screen "0887_Create Part Counter" 1280x800, template "Navigation"
   on GenerateScreen: SetTag("Create Part Counter Control", 1); SetTag("Create Part Counter Multiplexing Control", 0); function_b431313b("Part Counter Name", U 1, N)
   TextField "Text field_1" at 137,226 size 48x32; Text '1.'
      Visibility <- "Create Part Counter Control"
   TextField "Text field_2" at 137,266 size 48x32; Text '2.'
      Visibility <- "Create Part Counter Control"
   TextField "Text field_3" at 137,306 size 48x32; Text '3.'
      Visibility <- "Create Part Counter Control"
   TextField "Text field_4" at 137,346 size 48x32; Text '4.'
      Visibility <- "Create Part Counter Control"
   TextField "Text field_5" at 137,386 size 48x32; Text '5.'
      Visibility <- "Create Part Counter Control"
   TextField "Text field_6" at 137,426 size 48x32; Text '6.'
      Visibility <- "Create Part Counter Control"
   TextField "Text field_7" at 137,466 size 48x32; Text '7.'
      Visibility <- "Create Part Counter Control"
   TextField "Text field_8" at 137,506 size 48x32; Text '8.'
      Visibility <- "Create Part Counter Control"
   TextField "Text field_9" at 137,546 size 48x32; Text '9.'
      Visibility <- "Create Part Counter Control"
   TextField "Text field_10" at 137,586 size 48x32; Text '10.'
      Visibility <- "Create Part Counter Control"
   TextField "Text field_11" at 489,226 size 48x32; Text '11.'
      Visibility <- "Create Part Counter Control"
   TextField "Text field_12" at 489,266 size 48x32; Text '12.'
      Visibility <- "Create Part Counter Control"
   TextField "Text field_13" at 489,306 size 48x32; Text '13.'
      Visibility <- "Create Part Counter Control"
   TextField "Text field_14" at 489,346 size 48x32; Text '14.'
      Visibility <- "Create Part Counter Control"
   TextField "Text field_15" at 489,386 size 48x32; Text '15.'
      Visibility <- "Create Part Counter Control"
   TextField "Text field_16" at 489,426 size 48x32; Text '16.'
      Visibility <- "Create Part Counter Control"
   TextField "Text field_17" at 489,466 size 48x32; Text '17.'
      Visibility <- "Create Part Counter Control"
   TextField "Text field_18" at 489,506 size 48x32; Text '18.'
      Visibility <- "Create Part Counter Control"
   TextField "Text field_19" at 489,546 size 48x32; Text '19.'
      Visibility <- "Create Part Counter Control"
   TextField "Text field_20" at 489,586 size 48x32; Text '20.'
      Visibility <- "Create Part Counter Control"
   TextField "Text field_21" at 832,226 size 48x32; Text '21.'
      Visibility <- "Create Part Counter Control"
   TextField "Text field_22" at 832,266 size 48x32; Text '22.'
      Visibility <- "Create Part Counter Control"
   TextField "Text field_23" at 832,306 size 48x32; Text '23.'
      Visibility <- "Create Part Counter Control"
   TextField "Text field_24" at 832,346 size 48x32; Text '24.'
      Visibility <- "Create Part Counter Control"
   TextField "Text field_25" at 832,386 size 48x32; Text '25.'
      Visibility <- "Create Part Counter Control"
   TextField "Text field_26" at 832,426 size 48x32; Text '26.'
      Visibility <- "Create Part Counter Control"
   TextField "Text field_27" at 832,466 size 48x32; Text '27.'
      Visibility <- "Create Part Counter Control"
   TextField "Text field_28" at 832,506 size 48x32; Text '28.'
      Visibility <- "Create Part Counter Control"
   TextField "Text field_29" at 832,546 size 48x32; Text '29.'
      Visibility <- "Create Part Counter Control"
   TextField "Text field_30" at 832,586 size 48x32; Text '30.'
      Visibility <- "Create Part Counter Control"
   TextField "Text field_31" at 137,226 size 48x32; Text '31.'
      Visibility <- "Create Part Counter Control"
   TextField "Text field_32" at 137,266 size 48x32; Text '32.'
      Visibility <- "Create Part Counter Control"
   TextField "Text field_33" at 137,306 size 48x32; Text '33.'
      Visibility <- "Create Part Counter Control"
   TextField "Text field_34" at 137,346 size 48x32; Text '34.'
      Visibility <- "Create Part Counter Control"
   TextField "Text field_35" at 137,386 size 48x32; Text '35.'
      Visibility <- "Create Part Counter Control"
   TextField "Text field_36" at 137,426 size 48x32; Text '36.'
      Visibility <- "Create Part Counter Control"
   TextField "Text field_37" at 137,466 size 48x32; Text '37.'
      Visibility <- "Create Part Counter Control"
   TextField "Text field_38" at 137,506 size 48x32; Text '38.'
      Visibility <- "Create Part Counter Control"
   TextField "Text field_39" at 137,546 size 48x32; Text '39.'
      Visibility <- "Create Part Counter Control"
   TextField "Text field_40" at 137,586 size 48x32; Text '40.'
      Visibility <- "Create Part Counter Control"
   TextField "Text field_41" at 489,226 size 48x32; Text '41.'
      Visibility <- "Create Part Counter Control"
   TextField "Text field_42" at 489,266 size 48x32; Text '42.'
      Visibility <- "Create Part Counter Control"
   TextField "Text field_43" at 489,306 size 48x32; Text '43.'
      Visibility <- "Create Part Counter Control"
   TextField "Text field_44" at 489,346 size 48x32; Text '44.'
      Visibility <- "Create Part Counter Control"
   TextField "Text field_45" at 489,386 size 48x32; Text '45.'
      Visibility <- "Create Part Counter Control"
   TextField "Text field_46" at 489,426 size 48x32; Text '46.'
      Visibility <- "Create Part Counter Control"
   TextField "Text field_47" at 489,466 size 48x32; Text '47.'
      Visibility <- "Create Part Counter Control"
   TextField "Text field_48" at 489,506 size 48x32; Text '48.'
      Visibility <- "Create Part Counter Control"
   TextField "Text field_49" at 489,546 size 48x32; Text '49.'
      Visibility <- "Create Part Counter Control"
   TextField "Text field_50" at 489,586 size 48x32; Text '50.'
      Visibility <- "Create Part Counter Control"
   TextField "Text field_51" at 832,226 size 48x32; Text '51.'
      Visibility <- "Create Part Counter Control"
   TextField "Text field_52" at 832,266 size 48x32; Text '52.'
      Visibility <- "Create Part Counter Control"
   TextField "Text field_53" at 832,306 size 48x32; Text '53.'
      Visibility <- "Create Part Counter Control"
   TextField "Text field_54" at 832,346 size 48x32; Text '54.'
      Visibility <- "Create Part Counter Control"
   TextField "Text field_55" at 832,386 size 48x32; Text '55.'
      Visibility <- "Create Part Counter Control"
   TextField "Text field_56" at 832,426 size 48x32; Text '56.'
      Visibility <- "Create Part Counter Control"
   TextField "Text field_57" at 832,466 size 48x32; Text '57.'
      Visibility <- "Create Part Counter Control"
   TextField "Text field_58" at 832,506 size 48x32; Text '58.'
      Visibility <- "Create Part Counter Control"
   TextField "Text field_59" at 832,546 size 48x32; Text '59.'
      Visibility <- "Create Part Counter Control"
   TextField "Text field_60" at 832,586 size 48x32; Text '60.'
      Visibility <- "Create Part Counter Control"
   TextField "Text field_61" at 137,226 size 48x32; Text '61.'
      Visibility <- "Create Part Counter Control"
   TextField "Text field_62" at 137,266 size 48x32; Text '62.'
      Visibility <- "Create Part Counter Control"
   TextField "Text field_63" at 137,306 size 48x32; Text '63.'
      Visibility <- "Create Part Counter Control"
   TextField "Text field_64" at 137,346 size 48x32; Text '64.'
      Visibility <- "Create Part Counter Control"
   TextField "Text field_65" at 137,386 size 48x32; Text '65.'
      Visibility <- "Create Part Counter Control"
   TextField "Text field_66" at 137,426 size 48x32; Text '66.'
      Visibility <- "Create Part Counter Control"
   TextField "Text field_67" at 137,466 size 48x32; Text '67.'
      Visibility <- "Create Part Counter Control"
   TextField "Text field_68" at 137,506 size 48x32; Text '68.'
      Visibility <- "Create Part Counter Control"
   TextField "Text field_69" at 137,546 size 48x32; Text '69.'
      Visibility <- "Create Part Counter Control"
   TextField "Text field_70" at 137,586 size 48x32; Text '70.'
      Visibility <- "Create Part Counter Control"
   TextField "Text field_71" at 489,226 size 48x32; Text '71.'
      Visibility <- "Create Part Counter Control"
   TextField "Text field_72" at 489,266 size 48x32; Text '72.'
      Visibility <- "Create Part Counter Control"
   TextField "Text field_73" at 489,306 size 48x32; Text '73.'
      Visibility <- "Create Part Counter Control"
   TextField "Text field_74" at 489,346 size 48x32; Text '74.'
      Visibility <- "Create Part Counter Control"
   TextField "Text field_75" at 489,386 size 48x32; Text '75.'
      Visibility <- "Create Part Counter Control"
   TextField "Text field_76" at 489,426 size 48x32; Text '76.'
      Visibility <- "Create Part Counter Control"
   TextField "Text field_77" at 489,466 size 48x32; Text '77.'
      Visibility <- "Create Part Counter Control"
   TextField "Text field_78" at 489,506 size 48x32; Text '78.'
      Visibility <- "Create Part Counter Control"
   TextField "Text field_79" at 489,546 size 48x32; Text '79.'
      Visibility <- "Create Part Counter Control"
   TextField "Text field_80" at 489,586 size 48x32; Text '80.'
      Visibility <- "Create Part Counter Control"
   TextField "Text field_81" at 832,226 size 48x32; Text '81.'
      Visibility <- "Create Part Counter Control"
   TextField "Text field_82" at 832,266 size 48x32; Text '82.'
      Visibility <- "Create Part Counter Control"
   TextField "Text field_83" at 832,306 size 48x32; Text '83.'
      Visibility <- "Create Part Counter Control"
   TextField "Text field_84" at 832,346 size 48x32; Text '84.'
      Visibility <- "Create Part Counter Control"
   TextField "Text field_85" at 832,386 size 48x32; Text '85.'
      Visibility <- "Create Part Counter Control"
   TextField "Text field_86" at 832,426 size 48x32; Text '86.'
      Visibility <- "Create Part Counter Control"
   TextField "Text field_87" at 832,466 size 48x32; Text '87.'
      Visibility <- "Create Part Counter Control"
   TextField "Text field_88" at 832,506 size 48x32; Text '88.'
      Visibility <- "Create Part Counter Control"
   TextField "Text field_89" at 832,546 size 48x32; Text '89.'
      Visibility <- "Create Part Counter Control"
   TextField "Text field_90" at 832,586 size 48x32; Text '90.'
      Visibility <- "Create Part Counter Control"
   TextField "Text field_151" at 489,226 size 48x32; Text '101.'
      Visibility <- "Create Part Counter Control"
   TextField "Text field_152" at 489,266 size 48x32; Text '102.'
      Visibility <- "Create Part Counter Control"
   TextField "Text field_153" at 489,306 size 48x32; Text '103.'
      Visibility <- "Create Part Counter Control"
   TextField "Text field_154" at 489,346 size 48x32; Text '104.'
      Visibility <- "Create Part Counter Control"
   TextField "Text field_155" at 489,386 size 48x32; Text '105.'
      Visibility <- "Create Part Counter Control"
   TextField "Text field_156" at 489,426 size 48x32; Text '106.'
      Visibility <- "Create Part Counter Control"
   TextField "Text field_157" at 489,466 size 48x32; Text '107.'
      Visibility <- "Create Part Counter Control"
   TextField "Text field_158" at 489,506 size 48x32; Text '108.'
      Visibility <- "Create Part Counter Control"
   TextField "Text field_159" at 489,546 size 48x32; Text '109.'
      Visibility <- "Create Part Counter Control"
   TextField "Text field_160" at 489,586 size 48x32; Text '110.'
      Visibility <- "Create Part Counter Control"
   TextField "Text field_161" at 832,226 size 48x32; Text '111.'
      Visibility <- "Create Part Counter Control"
   TextField "Text field_162" at 832,266 size 48x32; Text '112.'
      Visibility <- "Create Part Counter Control"
   TextField "Text field_163" at 832,306 size 48x32; Text '113.'
      Visibility <- "Create Part Counter Control"
   TextField "Text field_164" at 832,346 size 48x32; Text '114.'
      Visibility <- "Create Part Counter Control"
   TextField "Text field_165" at 832,386 size 48x32; Text '115.'
      Visibility <- "Create Part Counter Control"
   TextField "Text field_166" at 832,426 size 48x32; Text '116.'
      Visibility <- "Create Part Counter Control"
   TextField "Text field_167" at 832,466 size 48x32; Text '117.'
      Visibility <- "Create Part Counter Control"
   TextField "Text field_168" at 832,506 size 48x32; Text '118.'
      Visibility <- "Create Part Counter Control"
   TextField "Text field_169" at 832,546 size 48x32; Text '119.'
      Visibility <- "Create Part Counter Control"
   TextField "Text field_170" at 832,586 size 48x32; Text '120.'
      Visibility <- "Create Part Counter Control"
   TextField "Text field_171" at 137,226 size 48x32; Text '91.'
      Visibility <- "Create Part Counter Control"
   TextField "Text field_172" at 137,266 size 48x32; Text '92.'
      Visibility <- "Create Part Counter Control"
   TextField "Text field_173" at 137,306 size 48x32; Text '93.'
      Visibility <- "Create Part Counter Control"
   TextField "Text field_174" at 137,346 size 48x32; Text '94.'
      Visibility <- "Create Part Counter Control"
   TextField "Text field_175" at 137,386 size 48x32; Text '95.'
      Visibility <- "Create Part Counter Control"
   TextField "Text field_176" at 137,426 size 48x32; Text '96.'
      Visibility <- "Create Part Counter Control"
   TextField "Text field_177" at 137,466 size 48x32; Text '97.'
      Visibility <- "Create Part Counter Control"
   TextField "Text field_178" at 137,506 size 48x32; Text '98.'
      Visibility <- "Create Part Counter Control"
   TextField "Text field_179" at 137,546 size 48x32; Text '99.'
      Visibility <- "Create Part Counter Control"
   TextField "Text field_180" at 137,586 size 48x32; Text '100.'
      Visibility <- "Create Part Counter Control"
   IOField "NamePart1" at 207,225 size 240x32; FormatPattern ????????????????????
      on OnFinishInput: SetTag("Create Part Counter Button Save", 1)
      ProcessValue <- "Part_Counter_Coloum_1"
   Button "Button_3" at 326,104 size 451x32; TextOff 'Create Part Counter'
   IOField "NamePart2" at 207,265 size 240x32; FormatPattern ????????????????????
      on OnFinishInput: SetTag("Create Part Counter Button Save", 1)
      ProcessValue <- "Part_Counter_Coloum_2"
   IOField "NamePart3" at 207,305 size 240x32; FormatPattern ????????????????????
      on OnFinishInput: SetTag("Create Part Counter Button Save", 1)
      ProcessValue <- "Part_Counter_Coloum_3"
   IOField "NamePart4" at 207,345 size 240x32; FormatPattern ????????????????????
      on OnFinishInput: SetTag("Create Part Counter Button Save", 1)
      ProcessValue <- "Part_Counter_Coloum_4"
   IOField "NamePart5" at 207,385 size 240x32; FormatPattern ????????????????????
      on OnFinishInput: SetTag("Create Part Counter Button Save", 1)
      ProcessValue <- "Part_Counter_Coloum_5"
   IOField "NamePart6" at 207,425 size 240x32; FormatPattern ????????????????????
      on OnFinishInput: SetTag("Create Part Counter Button Save", 1)
      ProcessValue <- "Part_Counter_Coloum_6"
   IOField "NamePart7" at 207,465 size 240x32; FormatPattern ????????????????????
      on OnFinishInput: SetTag("Create Part Counter Button Save", 1)
      ProcessValue <- "Part_Counter_Coloum_7"
   IOField "NamePart8" at 207,505 size 240x32; FormatPattern ????????????????????
      on OnFinishInput: SetTag("Create Part Counter Button Save", 1)
      ProcessValue <- "Part_Counter_Coloum_8"
   IOField "NamePart9" at 207,545 size 240x32; FormatPattern ????????????????????
      on OnFinishInput: SetTag("Create Part Counter Button Save", 1)
      ProcessValue <- "Part_Counter_Coloum_9"
   IOField "NamePart10" at 207,585 size 240x32; FormatPattern ????????????????????
      on OnFinishInput: SetTag("Create Part Counter Button Save", 1)
      ProcessValue <- "Part_Counter_Coloum_10"
   IOField "NamePart11" at 552,226 size 240x32; FormatPattern ????????????????????
      on OnFinishInput: SetTag("Create Part Counter Button Save", 1)
      ProcessValue <- "Part_Counter_Coloum_11"
   IOField "NamePart12" at 552,266 size 240x32; FormatPattern ????????????????????
      on OnFinishInput: SetTag("Create Part Counter Button Save", 1)
      ProcessValue <- "Part_Counter_Coloum_12"
   IOField "NamePart13" at 552,306 size 240x32; FormatPattern ????????????????????
      on OnFinishInput: SetTag("Create Part Counter Button Save", 1)
      ProcessValue <- "Part_Counter_Coloum_13"
   IOField "NamePart14" at 552,346 size 240x32; FormatPattern ????????????????????
      on OnFinishInput: SetTag("Create Part Counter Button Save", 1)
      ProcessValue <- "Part_Counter_Coloum_14"
   IOField "NamePart15" at 552,386 size 240x32; FormatPattern ????????????????????
      on OnFinishInput: SetTag("Create Part Counter Button Save", 1)
      ProcessValue <- "Part_Counter_Coloum_15"
   IOField "NamePart16" at 552,426 size 240x32; FormatPattern ????????????????????
      on OnFinishInput: SetTag("Create Part Counter Button Save", 1)
      ProcessValue <- "Part_Counter_Coloum_16"
   IOField "NamePart17" at 552,466 size 240x32; FormatPattern ????????????????????
      on OnFinishInput: SetTag("Create Part Counter Button Save", 1)
      ProcessValue <- "Part_Counter_Coloum_17"
   IOField "NamePart18" at 552,506 size 240x32; FormatPattern ????????????????????
      on OnFinishInput: SetTag("Create Part Counter Button Save", 1)
      ProcessValue <- "Part_Counter_Coloum_18"
   IOField "NamePart19" at 552,546 size 240x32; FormatPattern ????????????????????
      on OnFinishInput: SetTag("Create Part Counter Button Save", 1)
      ProcessValue <- "Part_Counter_Coloum_19"
   IOField "NamePart20" at 552,586 size 240x32; FormatPattern ????????????????????
      on OnFinishInput: SetTag("Create Part Counter Button Save", 1)
      ProcessValue <- "Part_Counter_Coloum_20"
   IOField "NamePart21" at 895,225 size 240x32; FormatPattern ????????????????????
      on OnFinishInput: SetTag("Create Part Counter Button Save", 1)
      ProcessValue <- "Part_Counter_Coloum_21"
   IOField "NamePart22" at 895,265 size 240x32; FormatPattern ????????????????????
      on OnFinishInput: SetTag("Create Part Counter Button Save", 1)
      ProcessValue <- "Part_Counter_Coloum_22"
   IOField "NamePart23" at 895,305 size 240x32; FormatPattern ????????????????????
      on OnFinishInput: SetTag("Create Part Counter Button Save", 1)
      ProcessValue <- "Part_Counter_Coloum_23"
   IOField "NamePart24" at 895,345 size 240x32; FormatPattern ????????????????????
      on OnFinishInput: SetTag("Create Part Counter Button Save", 1)
      ProcessValue <- "Part_Counter_Coloum_24"
   IOField "NamePart25" at 895,385 size 240x32; FormatPattern ????????????????????
      on OnFinishInput: SetTag("Create Part Counter Button Save", 1)
      ProcessValue <- "Part_Counter_Coloum_25"
   IOField "NamePart26" at 895,425 size 240x32; FormatPattern ????????????????????
      on OnFinishInput: SetTag("Create Part Counter Button Save", 1)
      ProcessValue <- "Part_Counter_Coloum_26"
   IOField "NamePart27" at 895,465 size 240x32; FormatPattern ????????????????????
      on OnFinishInput: SetTag("Create Part Counter Button Save", 1)
      ProcessValue <- "Part_Counter_Coloum_27"
   IOField "NamePart28" at 895,505 size 240x32; FormatPattern ????????????????????
      on OnFinishInput: SetTag("Create Part Counter Button Save", 1)
      ProcessValue <- "Part_Counter_Coloum_28"
   IOField "NamePart29" at 895,545 size 240x32; FormatPattern ????????????????????
      on OnFinishInput: SetTag("Create Part Counter Button Save", 1)
      ProcessValue <- "Part_Counter_Coloum_29"
   IOField "NamePart30" at 895,585 size 240x32; FormatPattern ????????????????????
      on OnFinishInput: SetTag("Create Part Counter Button Save", 1)
      ProcessValue <- "Part_Counter_Coloum_30"
   Button "Button_32" at 656,696 size 104x72; TextOff 'Text'; PictureOff "Tombol Increase"
      Visibility <- "Create Part Counter Control"
      on Click: function_dd21b452("Create Part Counter Control", 1); function_dd21b452("Create Part Counter Multiplexing Control", 1)
   Button "Button_33" at 464,696 size 104x72; TextOff 'Text'; PictureOff "Tombol Decrease"
      Visibility <- "Create Part Counter Control"
      on Click: function_b9b71300("Create Part Counter Control", 1); function_b9b71300("Create Part Counter Multiplexing Control", 1)
   Button "Button_34" at 976,696 size 104x72; TextOff 'Text'; PictureOff "Save_Icon"
      Visibility <- "Create Part Counter Button Save"
      on Click: SetTag("Create Part Counter Button Save", 0); function_f38ba6b2("Part Counter Name", U 1, 1, 1, N)

screen "0014_Network Setting" 1280x800, template "Navigation"
   Button "Button_3" at 326,99 size 451x32; TextOff 'Network Settings'
   TextField "Text field_1" at 260,370 size 180x27; Text 'Computer Name'
   IOField "I/O field_1" at 466,364 size 458x40; FormatPattern ????????????????????
      ProcessValue <- "Computer_Name"
   TextField "Text field_2" at 260,456 size 164x27; Text 'Enabled ordner'
   IOField "I/O field_2" at 466,450 size 458x40; FormatPattern ??????????
      ProcessValue <- "Ordner_Number"
   Button "Button_1" at 948,358 size 55x56; TextOff 'Text'
   Button "Button_2" at 948,429 size 55x56; TextOff 'Text'
   Button "Button_4" at 948,507 size 55x56; TextOff 'Text'

PopupScreen "Save" 350x130
   on GenerateScreen: SetBit("PopUp_Restrict")
   TextField "Text field_1" at 102,27 size 160x40; Text 'Text'
   GraphicView "Graphic view_1" at 19,28 size 47x40; Picture "Alarm Icon 1"
      Visibility <- "DB_MouldEditor_HMI_uData_sStatusBits"
   Button "Template_Button_24" at 158,90 size 45x30; TextOff 'Text'; PictureList "Check_Uncheck"; PictureOff "images (7)"
      ProcessValue <- "DB_MouldEditor_HMI_uData_arShotSet{3}_CPMoveAfterShot"
      on Click: SetBit("DB_MouldEditor_HMI_uData_sStatusBits_xDiscardChanges"); function_efd93a16("Save", 0, 0, 0, -1, 1); ResetBit("DB_MouldEditor_HMI_uData_sStatusBits_xValueChanged"); ResetBit("DB_MouldEditor_HMI_uData_sStatusBits_xFaultDeleteProgram"); ResetBit("DB_MouldEditor_HMI_uData_sStatusBits_xFaultValuesnotvalid"); ResetBit("PopUp_Restrict")
   Button "Template_Button_1" at 93,89 size 45x30; TextOff 'Text'; PictureList "Check_Uncheck"; PictureOff "_green_check.svg"
      ProcessValue <- "DB_MouldEditor_HMI_uData_arShotSet{3}_CPMoveAfterShot"
      on Click: SetBit("DB_MouldEditor_HMI_uData_sStatusBits_xSafeChanges"); SetBit("DB939_Tool_alloc_HMI_Delete_tool_in _all_allocations"); function_efd93a16("Save", 0, 0, -1, -1, 1); ResetBit("PopUp_Restrict")
   Button "Template_Button_2" at 222,91 size 45x30; TextOff 'TA'; PictureOff "Red_Checkmark"; PictureList "Check_Uncheck"
      ProcessValue <- "DB_MouldEditor_HMI_uData_arShotSet{3}_CPMoveAfterShot"
      on Click: ActivateScreen("0030_Tool Allocation", 0); ResetBit("DB_MouldEditor_HMI_uData_sStatusBits_xFaultDeleteProgram"); ResetBit("PopUp_Restrict")
      Visibility <- "DB_MouldEditor_HMI_uData_sStatusBits"

screen "0034_Robot" 1280x800, template "Navigation"
   on GenerateScreen: SetBit("DB1900_IF_Robots_Read"); SetBit("DB1901_Config_Robots_Read"); SetTag("Navigation_7", 6)
   Circle "Circle_1" at 166,243 size 21x21
      Appearance <- "DB1900_IF_Robots_State_Robots{0}_EmergencyStopReady"
   Button "b_Incress_Pump_Setting" at 784,104 size 46x32; TextOff 'Text'; PictureOff "right arrow"
      on Click: function_dd21b452("DB1900_IF_Robots_ReadWriteDeviceNo", 1)
   Button "b_Decress_Pump_Setting" at 273,104 size 46x32; TextOff 'Text'; PictureOff "left arrow"
      on Click: function_b9b71300("DB1900_IF_Robots_ReadWriteDeviceNo", 1)
   Circle "Circle_2" at 166,288 size 21x21
      Appearance <- "DB1900_IF_Robots_State_Robots{0}_AutomatcStopReady"
   Circle "Circle_3" at 166,333 size 21x21
      Appearance <- "DB1900_IF_Robots_State_Robots{0}_MaschineAuto"
   Circle "Circle_4" at 166,378 size 21x21
      Appearance <- "DB1900_IF_Robots_State_Robots{0}_MixingheadAuto"
   Circle "Circle_5" at 166,423 size 21x21
      Appearance <- "DB1900_IF_Robots_State_Robots{0}_Rob_in_Automatic"
   TextField "Text field_1" at 203,243 size 135x22; Text 'Control voltage'
   TextField "Text field_2" at 203,288 size 130x22; Text 'Automatic stop'
   TextField "Text field_3" at 203,333 size 121x22; Text 'OM Automatic'
   TextField "Text field_4" at 203,378 size 152x22; Text 'OM MH Automatic'
   TextField "Text field_5" at 203,423 size 175x22; Text 'OM Robot Automatic'
   Circle "Circle_6" at 493,243 size 21x21
      Appearance <- "DB1900_IF_Robots_State_Robots{0}_Rob_in_Home"
   Circle "Circle_7" at 495,333 size 21x21
      Appearance <- "DB1900_IF_Robots_State_Robots{0}_Rob_in_Cycle"
   TextField "Text field_6" at 224,472 size 186x22; Text 'Mould carrier number'
      Visibility <- "DB1900_IF_Robots_State_Robots{0}_TestShotRunning"
   TextField "Text field_7" at 226,510 size 143x22; Text 'Program number'
      Visibility <- "DB1900_IF_Robots_State_Robots{0}_TestShotRunning"
   IOField "I/O field_1" at 420,470 size 60x24; FormatPattern 9999
      Visibility <- "DB1900_IF_Robots_State_Robots{0}_TestShotRunning"
      ProcessValue <- "DB1900_IF_Robots_State_Robots{0}_Rob_MC_No"
   IOField "I/O field_2" at 420,508 size 60x24; FormatPattern 9999
      Visibility <- "DB1900_IF_Robots_State_Robots{0}_TestShotRunning"
      ProcessValue <- "DB1900_IF_Robots_State_Robots{0}_Rob_Prog_No"
   GraphicView "Graphic view_1" at 650,602 size 68x182; Picture "robo_2"
      Visibility <- "DB1901_Config_Robots_Config_Robots{0}_With_Cleaning"
   GraphicView "ABB ROBOT" at 578,227 size 198x244; Picture "ABB Robot"
      Visibility <- "DB1901_Config_Robots_Config_Robots{0}_Type_ABB"
   GraphicView "KUKA ROBOT" at 578,227 size 198x244; Picture "Kuka Robot"
      Visibility <- "DB1901_Config_Robots_Config_Robots{0}_Type_Kuka"
   GraphicView "MOTOMAN ROBOT" at 578,227 size 198x244; Picture "Motoman Robot"
      Visibility <- "DB1901_Config_Robots_Config_Robots{0}_Type_Motoman"
   GraphicView "FANUC ROBOT" at 578,227 size 198x244; Picture "Fanuc Robot"
      Visibility <- "DB1901_Config_Robots_Config_Robots{0}_Type_Fanuc"
   Button "Button_5" at 797,235 size 81x116; TextOff 'Text'
   GraphicView "Graphic view_5" at 809,300 size 56x45; Picture "settingrobot"
   Rectangle "Rectangle_6" at 806,243 size 64x56
      Appearance <- "DB1900_IF_Robots_Switch_Robots{0}_StateMaintPos"
   GraphicIOField "Graphic I/O field_5" at 814,246 size 48x48; PictureList "ON_OFF_SWITCH"
      ProcessValue <- "DB1900_IF_Robots_Switch_Robots{0}_SwitchMaintPosON_OFF"
   Button "Button_22" at 793,227 size 88x128; TextOff 'Text'
      on Click: InvertBit("DB1900_IF_Robots_Switch_Robots{0}_SwitchMaintPosON_OFF")
   Button "Button_3" at 892,235 size 81x116; TextOff 'Text'
   GraphicView "Graphic view_2" at 911,300 size 56x44; Picture "settingrobot"
   Rectangle "Rectangle_1" at 901,243 size 64x56
      Appearance <- "DB1900_IF_Robots_Switch_Robots{0}_StateMaintPos_2"
   GraphicIOField "Graphic I/O field_1" at 909,246 size 48x48; PictureList "ON_OFF_SWITCH"
      ProcessValue <- "DB1900_IF_Robots_Switch_Robots{0}_SwitchMaintPos_2ON_OFF"
   Button "Button_6" at 987,235 size 81x116; TextOff 'Text'
      Visibility <- "DB1901_Config_Robots_Config_Robots{0}_With_Wet_Cleaning_LFI"
   GraphicView "Graphic view_3" at 999,302 size 56x43; Picture "LFI"
      Visibility <- "DB1901_Config_Robots_Config_Robots{0}_With_Wet_Cleaning_LFI"
   Rectangle "Rectangle_3" at 996,243 size 64x56
      Appearance <- "DB1900_IF_Robots_Switch_Robots{0}_StateCleaning"
      Visibility <- "DB1901_Config_Robots_Config_Robots{0}_With_Wet_Cleaning_LFI"
   Button "Button_4" at 888,227 size 88x128; TextOff 'Text'
      on Click: InvertBit("DB1900_IF_Robots_Switch_Robots{0}_SwitchMaintPos_2ON_OFF")
   GraphicIOField "Graphic I/O field_2" at 1004,246 size 48x48; PictureList "ON_OFF_SWITCH"
      ProcessValue <- "DB1900_IF_Robots_Switch_Robots{0}_SwitchCleaningON_OFF"
      Visibility <- "DB1901_Config_Robots_Config_Robots{0}_With_Wet_Cleaning_LFI"
   Button "Button_7" at 983,227 size 88x128; TextOff 'Text'
      on Click: InvertBit("DB1900_IF_Robots_Switch_Robots{0}_SwitchCleaningON_OFF")
      Visibility <- "DB1901_Config_Robots_Config_Robots{0}_With_Wet_Cleaning_LFI"
   Button "Button_8" at 798,386 size 81x116; TextOff 'Text'
      Visibility <- "DB1901_Config_Robots_Config_Robots{0}_With_Cleaning"
   GraphicView "Graphic view_4" at 816,451 size 42x43; Picture "brush"
      Visibility <- "DB1901_Config_Robots_Config_Robots{0}_With_Cleaning"
   Rectangle "Rectangle_4" at 807,394 size 64x56
      Appearance <- "DB1900_IF_Robots_Switch_Robots{0}_StateBrush"
      Visibility <- "DB1901_Config_Robots_Config_Robots{0}_With_Cleaning"
   GraphicIOField "Graphic I/O field_3" at 815,397 size 48x48; PictureList "ON_OFF_SWITCH"
      ProcessValue <- "DB1900_IF_Robots_Switch_Robots{0}_SwitchBrushON_OFF"
      Visibility <- "DB1901_Config_Robots_Config_Robots{0}_With_Cleaning"
   Button "Button_9" at 794,378 size 88x128; TextOff 'Text'
      on Click: InvertBit("DB1900_IF_Robots_Switch_Robots{0}_SwitchBrushON_OFF")
      Visibility <- "DB1901_Config_Robots_Config_Robots{0}_With_Cleaning"
   Button "Button_10" at 893,386 size 81x116; TextOff 'Text'
      Visibility <- "DB1901_Config_Robots_Config_Robots{0}_With_Synchronisation"
   GraphicView "Graphic view_6" at 905,451 size 56x48; Picture "circ_robot"
      Visibility <- "DB1901_Config_Robots_Config_Robots{0}_With_Synchronisation"
   Rectangle "Rectangle_5" at 902,394 size 64x56
      Appearance <- "DB1900_IF_Robots_Switch_Robots{0}_StateSync"
      Visibility <- "DB1901_Config_Robots_Config_Robots{0}_With_Synchronisation"
   GraphicIOField "Graphic I/O field_4" at 910,397 size 48x48; PictureList "ON_OFF_SWITCH"
      ProcessValue <- "DB1900_IF_Robots_Switch_Robots{0}_SwitchSyncON_OFF"
      Visibility <- "DB1901_Config_Robots_Config_Robots{0}_With_Synchronisation"
   Button "Button_11" at 889,378 size 88x128; TextOff 'Text'
      on Click: InvertBit("DB1900_IF_Robots_Switch_Robots{0}_SwitchSyncON_OFF")
      Visibility <- "DB1901_Config_Robots_Config_Robots{0}_With_Synchronisation"
   Button "Button_12" at 988,386 size 81x116; TextOff 'Text'
      Visibility <- "DB1901_Config_Robots_Config_Robots{0}_With_Air_Cleaner"
   GraphicView "Graphic view_7" at 1000,447 size 56x48; Picture "CleaningPiston"
      Visibility <- "DB1901_Config_Robots_Config_Robots{0}_With_Air_Cleaner"
   Rectangle "Rectangle_7" at 997,394 size 64x56
      Appearance <- "DB1900_IF_Robots_Switch_Robots{0}_StateAirCleaning"
      Visibility <- "DB1901_Config_Robots_Config_Robots{0}_With_Air_Cleaner"
   GraphicIOField "Graphic I/O field_6" at 1005,397 size 48x48; PictureList "ON_OFF_SWITCH"
      ProcessValue <- "DB1900_IF_Robots_Switch_Robots{0}_SwitchAirCleaningON_OFF"
      Visibility <- "DB1901_Config_Robots_Config_Robots{0}_With_Air_Cleaner"
   Button "Button_13" at 984,378 size 88x128; TextOff 'Text'
      on Click: InvertBit("DB1900_IF_Robots_Switch_Robots{0}_SwitchAirCleaningON_OFF")
      Visibility <- "DB1901_Config_Robots_Config_Robots{0}_With_Air_Cleaner"
   Button "Button_14" at 1082,387 size 81x116; TextOff 'Text'
      Visibility <- "DB1901_Config_Robots_Config_Robots{0}_With_Air_Cleaner"
   GraphicView "Graphic view_8" at 1094,448 size 56x48; Picture "CleaningPiston"
      Visibility <- "DB1901_Config_Robots_Config_Robots{0}_With_Air_Cleaner"
   Rectangle "Rectangle_8" at 1091,395 size 64x56
      Appearance <- "DB1900_IF_Robots_Switch_Robots{0}_StateAirCleaningManual"
      Visibility <- "DB1901_Config_Robots_Config_Robots{0}_With_Air_Cleaner"
   GraphicIOField "Graphic I/O field_7" at 1099,398 size 48x48; PictureList "ON_OFF_SWITCH"
      ProcessValue <- "DB1900_IF_Robots_Switch_Robots{0}_SwitchAirCleaningManON_OFF"
      Visibility <- "DB1901_Config_Robots_Config_Robots{0}_With_Air_Cleaner"
   Button "Button_15" at 1078,379 size 88x128; TextOff 'Text'
      on Click: InvertBit("DB1900_IF_Robots_Switch_Robots{0}_SwitchAirCleaningManON_OFF")
      Visibility <- "DB1901_Config_Robots_Config_Robots{0}_With_Air_Cleaner"
   GraphicView "Graphic view_9" at 422,223 size 64x61; Picture "Graphic_5"
   GraphicView "Graphic view_10" at 422,313 size 64x61; Picture "Graphic_6"
   Button "Button_16" at 177,170 size 960x37; TextOff '----------------------------------------------'
   GraphicView "Graphic view_11" at 409,579 size 138x204; Picture "IR Station"
      Visibility <- "DB1901_Config_Robots_Config_Robots{0}_With_IR_Station"
   GraphicView "Graphic view_12" at 410,579 size 138x204; Picture "LFI"
      Visibility <- "DB1901_Config_Robots_Config_Robots{0}_With_Wet_Cleaning_LFI"
   GraphicView "Graphic view_13" at 170,588 size 138x204; Picture "spare"
      Visibility <- "DB1901_Config_Robots_Config_Robots{0}_With_Belt_Filter"
   GraphicView "Graphic view_14" at 170,566 size 328x225; Picture "Spray Clean"
      Visibility <- "DB1901_Config_Robots_Config_Robots{0}_With_Wet_Cleaning_Spray"
   GraphicView "Graphic view_15" at 570,602 size 68x182; Picture "robo_2"
      Visibility <- "DB1901_Config_Robots_Config_Robots{0}_With_Brush_Station"
   TextField "Text field_8" at 897,302 size 56x29; Text '2.'
   SymbolicIOField "Symbolic I/O field_1" at 326,104 size 451x32; TextOff '0'; TextOn '1'; TextList "Robot_name"
      ProcessValue <- "DB1900_IF_Robots_ReadWriteDeviceNo"